HMI tags "DB_SDC_GLOBAL"
   "DB_SDC_GLOBAL_LIMITS[2].RAPID_SLOW" : Int = PLC DB_SDC_GLOBAL.LIMITS[2].RAPID_SLOW AT %DB3700.DBW512, 1 s   // Umstellung Begrenzung auf Abstand (mm), Einschränkung / Changeover limit of distance (mm), limitation
   "DB_SDC_GLOBAL_SYNCH[15].K" : Real = PLC DB_SDC_GLOBAL.SYNCH[15].K AT %DB3700.DBD426, 1 s   // erreichen von Synchron Faktor / gain for Synchron Faktor
   "DB_SDC_GLOBAL_SYNCH[15].SET_DIST" : Int = PLC DB_SDC_GLOBAL.SYNCH[15].SET_DIST AT %DB3700.DBW420, 1 s   // Set point value: distance (mm)
   "DB_SDC_GLOBAL_LIMITS[6].RAPID_SLOW" : Int = PLC DB_SDC_GLOBAL.LIMITS[6].RAPID_SLOW AT %DB3700.DBW536, 1 s   // Umstellung Begrenzung auf Abstand (mm), Einschränkung / Changeover limit of distance (mm), limitation
   "DB_SDC_GLOBAL_SYNCH[11].HYST" : Int = PLC DB_SDC_GLOBAL.SYNCH[11].HYST AT %DB3700.DBW352, 1 s   // IO Hysterese
   "DB_SDC_GLOBAL_SYNCH[6].MIN_FAKT" : Real = PLC DB_SDC_GLOBAL.SYNCH[6].MIN_FAKT AT %DB3700.DBD272, 1 s   // Faktor für minimale Synchronisiergeschwindigkeit / Faktor Speed for Synchron MIN
   "DB_SDC_GLOBAL_MIN_DIST_EMS[13]" : Int = PLC DB_SDC_GLOBAL.MIN_DIST_EMS[13] AT %DB3700.DBW126, 1 s   // minimum distance
   "DB_SDC_GLOBAL_SYNCH[8].MIN_FAKT" : Real = PLC DB_SDC_GLOBAL.SYNCH[8].MIN_FAKT AT %DB3700.DBD308, 1 s   // Faktor für minimale Synchronisiergeschwindigkeit / Faktor Speed for Synchron MIN
   "DB_SDC_GLOBAL_SYNCH[10].MIN_FAKT" : Real = PLC DB_SDC_GLOBAL.SYNCH[10].MIN_FAKT AT %DB3700.DBD344, 1 s   // Faktor für minimale Synchronisiergeschwindigkeit / Faktor Speed for Synchron MIN
   "DB_SDC_GLOBAL_SYNCH[6].SET_DIST" : Int = PLC DB_SDC_GLOBAL.SYNCH[6].SET_DIST AT %DB3700.DBW258, 1 s   // Set point value: distance (mm)
   "DB_SDC_GLOBAL_SYNCH[11].MAX_FAKT" : Real = PLC DB_SDC_GLOBAL.SYNCH[11].MAX_FAKT AT %DB3700.DBD358, 1 s   // Faktor für maximale Synchronisiergeschwindigkeit / Faktor Speed for Synchron MAX
   "DB_SDC_GLOBAL_SYNCH[9].SET_DIST" : Int = PLC DB_SDC_GLOBAL.SYNCH[9].SET_DIST AT %DB3700.DBW312, 1 s   // Set point value: distance (mm)
   "DB_SDC_GLOBAL_SYNCH[11].MIN_FAKT" : Real = PLC DB_SDC_GLOBAL.SYNCH[11].MIN_FAKT AT %DB3700.DBD362, 1 s   // Faktor für minimale Synchronisiergeschwindigkeit / Faktor Speed for Synchron MIN
   "DB_SDC_GLOBAL_MAN_V_1" : DInt = PLC DB_SDC_GLOBAL.MAN_V_1 AT %DB3700.DBD30, 1 s   // manual mode, set value: drive speed (mm/min)
   "DB_SDC_GLOBAL_LIMITS[5].RAPID_SLOW" : Int = PLC DB_SDC_GLOBAL.LIMITS[5].RAPID_SLOW AT %DB3700.DBW530, 1 s   // Umstellung Begrenzung auf Abstand (mm), Einschränkung / Changeover limit of distance (mm), limitation
   "DB_SDC_GLOBAL_SYNCH[13].MIN_FAKT" : Real = PLC DB_SDC_GLOBAL.SYNCH[13].MIN_FAKT AT %DB3700.DBD398, 1 s   // Faktor für minimale Synchronisiergeschwindigkeit / Faktor Speed for Synchron MIN
   "DB_SDC_GLOBAL_SYNCH[10].SET_DIST" : Int = PLC DB_SDC_GLOBAL.SYNCH[10].SET_DIST AT %DB3700.DBW330, 1 s   // Set point value: distance (mm)
   "DB_SDC_GLOBAL_SYNCH[9].HYST" : Int = PLC DB_SDC_GLOBAL.SYNCH[9].HYST AT %DB3700.DBW316, 1 s   // IO Hysterese
   "DB_SDC_GLOBAL_SYNCH[13].MAX_FAKT" : Real = PLC DB_SDC_GLOBAL.SYNCH[13].MAX_FAKT AT %DB3700.DBD394, 1 s   // Faktor für maximale Synchronisiergeschwindigkeit / Faktor Speed for Synchron MAX
   "DB_SDC_GLOBAL_LIMITS[11].RAPID_SLOW" : Int = PLC DB_SDC_GLOBAL.LIMITS[11].RAPID_SLOW AT %DB3700.DBW566, 1 s   // Umstellung Begrenzung auf Abstand (mm), Einschränkung / Changeover limit of distance (mm), limitation
   "DB_SDC_GLOBAL_SYNCH[3].MIN_FAKT" : Real = PLC DB_SDC_GLOBAL.SYNCH[3].MIN_FAKT AT %DB3700.DBD218, 1 s   // Faktor für minimale Synchronisiergeschwindigkeit / Faktor Speed for Synchron MIN
   "DB_SDC_GLOBAL_SYNCH[7].K" : Real = PLC DB_SDC_GLOBAL.SYNCH[7].K AT %DB3700.DBD282, 1 s   // erreichen von Synchron Faktor / gain for Synchron Faktor
   "DB_SDC_GLOBAL_SYNCH[2].SYNCH_DIST" : Int = PLC DB_SDC_GLOBAL.SYNCH[2].SYNCH_DIST AT %DB3700.DBW188, 1 s   // Start synchron distance value: distance (mm)
   "DB_SDC_GLOBAL_SYNCH[14].SYNCH_DIST" : Int = PLC DB_SDC_GLOBAL.SYNCH[14].SYNCH_DIST AT %DB3700.DBW404, 1 s   // Start synchron distance value: distance (mm)
   "DB_SDC_GLOBAL_MIN_DIST_EMS[8]" : Int = PLC DB_SDC_GLOBAL.MIN_DIST_EMS[8] AT %DB3700.DBW116, 1 s   // minimum distance
   "DB_SDC_GLOBAL_MIN_DIST_EMS[0]" : Int = PLC DB_SDC_GLOBAL.MIN_DIST_EMS[0] AT %DB3700.DBW100, 1 s   // minimum distance
   "DB_SDC_GLOBAL_SYNCH[14].K" : Real = PLC DB_SDC_GLOBAL.SYNCH[14].K AT %DB3700.DBD408, 1 s   // erreichen von Synchron Faktor / gain for Synchron Faktor
   "DB_SDC_GLOBAL_LIMITS[1].RAPID_SLOW" : Int = PLC DB_SDC_GLOBAL.LIMITS[1].RAPID_SLOW AT %DB3700.DBW506, 1 s   // Umstellung Begrenzung auf Abstand (mm), Einschränkung / Changeover limit of distance (mm), limitation
   "DB_SDC_GLOBAL_LIMITS[14].SLOW_SPEED_FAKT" : Real = PLC DB_SDC_GLOBAL.LIMITS[14].SLOW_SPEED_FAKT AT %DB3700.DBD586, 1 s   // Faktor Geschwindigkeit für langsame Drehzahl / Faktor Speed for Slow Speed
   "DB_SDC_GLOBAL_SYNCH[14].SET_DIST" : Int = PLC DB_SDC_GLOBAL.SYNCH[14].SET_DIST AT %DB3700.DBW402, 1 s   // Set point value: distance (mm)
   "DB_SDC_GLOBAL_SYNCH[15].SYNCH_DIST" : Int = PLC DB_SDC_GLOBAL.SYNCH[15].SYNCH_DIST AT %DB3700.DBW422, 1 s   // Start synchron distance value: distance (mm)
   "DB_SDC_GLOBAL_SYNCH[4].MAX_FAKT" : Real = PLC DB_SDC_GLOBAL.SYNCH[4].MAX_FAKT AT %DB3700.DBD232, 1 s   // Faktor für maximale Synchronisiergeschwindigkeit / Faktor Speed for Synchron MAX
   "DB_SDC_GLOBAL_SYNCH[2].HYST" : Int = PLC DB_SDC_GLOBAL.SYNCH[2].HYST AT %DB3700.DBW190, 1 s   // IO Hysterese
   "DB_SDC_GLOBAL_MIN_DIST_EMS[6]" : Int = PLC DB_SDC_GLOBAL.MIN_DIST_EMS[6] AT %DB3700.DBW112, 1 s   // minimum distance
   "DB_SDC_GLOBAL_SYNCH[0].HYST" : Int = PLC DB_SDC_GLOBAL.SYNCH[0].HYST AT %DB3700.DBW154, 1 s   // IO Hysterese
   "DB_SDC_GLOBAL_MIN_DIST_EMS[2]" : Int = PLC DB_SDC_GLOBAL.MIN_DIST_EMS[2] AT %DB3700.DBW104, 1 s   // minimum distance
   "DB_SDC_GLOBAL_MIN_DIST_EMS[12]" : Int = PLC DB_SDC_GLOBAL.MIN_DIST_EMS[12] AT %DB3700.DBW124, 1 s   // minimum distance
   "DB_SDC_GLOBAL_LIMITS[15].RAPID_SLOW" : Int = PLC DB_SDC_GLOBAL.LIMITS[15].RAPID_SLOW AT %DB3700.DBW590, 1 s   // Umstellung Begrenzung auf Abstand (mm), Einschränkung / Changeover limit of distance (mm), limitation
   "DB_SDC_GLOBAL_LIMITS[2].SLOW_SPEED_FAKT" : Real = PLC DB_SDC_GLOBAL.LIMITS[2].SLOW_SPEED_FAKT AT %DB3700.DBD514, 1 s   // Faktor Geschwindigkeit für langsame Drehzahl / Faktor Speed for Slow Speed
   "DB_SDC_GLOBAL_SYNCH[8].SET_DIST" : Int = PLC DB_SDC_GLOBAL.SYNCH[8].SET_DIST AT %DB3700.DBW294, 1 s   // Set point value: distance (mm)
   "DB_SDC_GLOBAL_min_barcode_mm" : DInt = PLC DB_SDC_GLOBAL.min_barcode_mm AT %DB3700.DBD6, 1 s   // Lower limit, bar code value
   "DB_SDC_GLOBAL_LIMITS[13].SLOW_SPEED_FAKT" : Real = PLC DB_SDC_GLOBAL.LIMITS[13].SLOW_SPEED_FAKT AT %DB3700.DBD580, 1 s   // Faktor Geschwindigkeit für langsame Drehzahl / Faktor Speed for Slow Speed
   "DB_SDC_GLOBAL_LIMITS[9].SLOW_SPEED_FAKT" : Real = PLC DB_SDC_GLOBAL.LIMITS[9].SLOW_SPEED_FAKT AT %DB3700.DBD556, 1 s   // Faktor Geschwindigkeit für langsame Drehzahl / Faktor Speed for Slow Speed
   "DB_SDC_GLOBAL_MIN_DIST_EMS[3]" : Int = PLC DB_SDC_GLOBAL.MIN_DIST_EMS[3] AT %DB3700.DBW106, 1 s   // minimum distance
   "DB_SDC_GLOBAL_SYNCH[4].SET_DIST" : Int = PLC DB_SDC_GLOBAL.SYNCH[4].SET_DIST AT %DB3700.DBW222, 1 s   // Set point value: distance (mm)
   "DB_SDC_GLOBAL_MAN_V_2" : DInt = PLC DB_SDC_GLOBAL.MAN_V_2 AT %DB3700.DBD34, 1 s   // manual mode, set value: drive speed (mm/min)
   "DB_SDC_GLOBAL_SYNCH[6].K" : Real = PLC DB_SDC_GLOBAL.SYNCH[6].K AT %DB3700.DBD264, 1 s   // erreichen von Synchron Faktor / gain for Synchron Faktor
   "DB_SDC_GLOBAL_SYNCH[2].K" : Real = PLC DB_SDC_GLOBAL.SYNCH[2].K AT %DB3700.DBD192, 1 s   // erreichen von Synchron Faktor / gain for Synchron Faktor
   "DB_SDC_GLOBAL_SYNCH[4].MIN_FAKT" : Real = PLC DB_SDC_GLOBAL.SYNCH[4].MIN_FAKT AT %DB3700.DBD236, 1 s   // Faktor für minimale Synchronisiergeschwindigkeit / Faktor Speed for Synchron MIN
   "DB_SDC_GLOBAL_SYNCH[6].SYNCH_DIST" : Int = PLC DB_SDC_GLOBAL.SYNCH[6].SYNCH_DIST AT %DB3700.DBW260, 1 s   // Start synchron distance value: distance (mm)
   "DB_SDC_GLOBAL_LIMITS[8].RAPID_SLOW" : Int = PLC DB_SDC_GLOBAL.LIMITS[8].RAPID_SLOW AT %DB3700.DBW548, 1 s   // Umstellung Begrenzung auf Abstand (mm), Einschränkung / Changeover limit of distance (mm), limitation
   "DB_SDC_GLOBAL_SYNCH[11].SET_DIST" : Int = PLC DB_SDC_GLOBAL.SYNCH[11].SET_DIST AT %DB3700.DBW348, 1 s   // Set point value: distance (mm)
   "DB_SDC_GLOBAL_SYNCH[15].HYST" : Int = PLC DB_SDC_GLOBAL.SYNCH[15].HYST AT %DB3700.DBW424, 1 s   // IO Hysterese
   "DB_SDC_GLOBAL_SYNCH[13].HYST" : Int = PLC DB_SDC_ERRORS_STAT.ER_AKT[50].ER_STAT[2].ERROR AT %DB3700.DBW388, 1 s   // IO Hysterese
   "DB_SDC_GLOBAL_SYNCH[5].MAX_FAKT" : Real = PLC DB_SDC_GLOBAL.SYNCH[5].MAX_FAKT AT %DB3700.DBD250, 1 s   // Faktor für maximale Synchronisiergeschwindigkeit / Faktor Speed for Synchron MAX
   "DB_SDC_GLOBAL_EMS_ID_MIN" : Int = PLC DB_SDC_GLOBAL.EMS_ID_MIN AT %DB3700.DBW2, 1 s   // Minimum EMS ID
   "DB_SDC_GLOBAL_SYNCH[5].K" : Real = PLC DB_SDC_GLOBAL.SYNCH[5].K AT %DB3700.DBD246, 1 s   // erreichen von Synchron Faktor / gain for Synchron Faktor
   "DB_SDC_GLOBAL_SYNCH[5].SET_DIST" : Int = PLC DB_SDC_GLOBAL.SYNCH[5].SET_DIST AT %DB3700.DBW240, 1 s   // Set point value: distance (mm)
   "DB_SDC_GLOBAL_SYNCH[0].SYNCH_DIST" : Int = PLC DB_SDC_GLOBAL.SYNCH[0].SYNCH_DIST AT %DB3700.DBW152, 1 s   // Start synchron distance value: distance (mm)
   "DB_SDC_GLOBAL_MIN_DIST_EMS[1]" : Int = PLC DB_SDC_GLOBAL.MIN_DIST_EMS[1] AT %DB3700.DBW102, 1 s   // minimum distance
   "DB_SDC_GLOBAL_SEK_MIN" : Int = PLC DB_SDC_GLOBAL.SEK_MIN AT %DB3700.DBW22, 1 s   // Erste Abschnitt Nummer / first section number
   "DB_SDC_GLOBAL_SYNCH[2].MAX_FAKT" : Real = PLC DB_SDC_GLOBAL.SYNCH[2].MAX_FAKT AT %DB3700.DBD196, 1 s   // Faktor für maximale Synchronisiergeschwindigkeit / Faktor Speed for Synchron MAX
   "DB_SDC_GLOBAL_SYNCH[1].MIN_FAKT" : Real = PLC DB_SDC_GLOBAL.SYNCH[1].MIN_FAKT AT %DB3700.DBD182, 1 s   // Faktor für minimale Synchronisiergeschwindigkeit / Faktor Speed for Synchron MIN
   "DB_SDC_GLOBAL_SYNCH[2].MIN_FAKT" : Real = PLC DB_SDC_GLOBAL.SYNCH[2].MIN_FAKT AT %DB3700.DBD200, 1 s   // Faktor für minimale Synchronisiergeschwindigkeit / Faktor Speed for Synchron MIN
   "DB_SDC_GLOBAL_LIMITS[10].RAPID_SLOW" : Int = PLC DB_SDC_GLOBAL.LIMITS[10].RAPID_SLOW AT %DB3700.DBW560, 1 s   // Umstellung Begrenzung auf Abstand (mm), Einschränkung / Changeover limit of distance (mm), limitation
   "DB_SDC_GLOBAL_SYNCH[6].MAX_FAKT" : Real = PLC DB_SDC_GLOBAL.SYNCH[6].MAX_FAKT AT %DB3700.DBD268, 1 s   // Faktor für maximale Synchronisiergeschwindigkeit / Faktor Speed for Synchron MAX
   "DB_SDC_GLOBAL_SYNCH[10].K" : Real = PLC DB_SDC_GLOBAL.SYNCH[10].K AT %DB3700.DBD336, 1 s   // erreichen von Synchron Faktor / gain for Synchron Faktor
   "DB_SDC_GLOBAL_END_COURSE" : DInt = PLC DB_SDC_GLOBAL.END_COURSE AT %DB3700.DBD18, 1 s   // Ende Barcodewert vom Kurs / End Barcodevalue of Course
   "DB_SDC_GLOBAL_SYNCH[1].SYNCH_DIST" : Int = PLC DB_SDC_GLOBAL.SYNCH[1].SYNCH_DIST AT %DB3700.DBW170, 1 s   // Start synchron distance value: distance (mm)
   "DB_SDC_GLOBAL_LIMITS[1].SLOW_SPEED_FAKT" : Real = PLC DB_SDC_GLOBAL.LIMITS[1].SLOW_SPEED_FAKT AT %DB3700.DBD508, 1 s   // Faktor Geschwindigkeit für langsame Drehzahl / Faktor Speed for Slow Speed
   "DB_SDC_GLOBAL_SYNCH[11].SYNCH_DIST" : Int = PLC DB_SDC_GLOBAL.SYNCH[11].SYNCH_DIST AT %DB3700.DBW350, 1 s   // Start synchron distance value: distance (mm)
   "DB_SDC_GLOBAL_SYNCH[12].HYST" : Int = PLC DB_SDC_GLOBAL.SYNCH[12].HYST AT %DB3700.DBW370, 1 s   // IO Hysterese
   "DB_SDC_GLOBAL_LIMITS[0].RAPID_SLOW" : Int = PLC DB_SDC_GLOBAL.LIMITS[0].RAPID_SLOW AT %DB3700.DBW500, 1 s   // Umstellung Begrenzung auf Abstand (mm), Einschränkung / Changeover limit of distance (mm), limitation
   "DB_SDC_GLOBAL_SYNCH[15].MIN_FAKT" : Real = PLC DB_SDC_GLOBAL.SYNCH[15].MIN_FAKT AT %DB3700.DBD434, 1 s   // Faktor für minimale Synchronisiergeschwindigkeit / Faktor Speed for Synchron MIN
   "DB_SDC_GLOBAL_LIMITS[11].SLOW_SPEED_FAKT" : Real = PLC DB_SDC_GLOBAL.LIMITS[11].SLOW_SPEED_FAKT AT %DB3700.DBD568, 1 s   // Faktor Geschwindigkeit für langsame Drehzahl / Faktor Speed for Slow Speed
   "DB_SDC_GLOBAL_LIMITS[6].SLOW_SPEED_FAKT" : Real = PLC DB_SDC_GLOBAL.LIMITS[6].SLOW_SPEED_FAKT AT %DB3700.DBD538, 1 s   // Faktor Geschwindigkeit für langsame Drehzahl / Faktor Speed for Slow Speed
   "DB_SDC_GLOBAL_SYNCH[3].SYNCH_DIST" : Int = PLC DB_SDC_GLOBAL.SYNCH[3].SYNCH_DIST AT %DB3700.DBW206, 1 s   // Start synchron distance value: distance (mm)
   "DB_SDC_GLOBAL_MIN_DIST_EMS[11]" : Int = PLC DB_SDC_GLOBAL.MIN_DIST_EMS[11] AT %DB3700.DBW122, 1 s   // minimum distance
   "DB_SDC_GLOBAL_SYNCH[9].MAX_FAKT" : Real = PLC DB_SDC_GLOBAL.SYNCH[9].MAX_FAKT AT %DB3700.DBD322, 1 s   // Faktor für maximale Synchronisiergeschwindigkeit / Faktor Speed for Synchron MAX
   "DB_SDC_GLOBAL_MIN_DIST_EMS[9]" : Int = PLC DB_SDC_GLOBAL.MIN_DIST_EMS[9] AT %DB3700.DBW118, 1 s   // minimum distance
   "DB_SDC_GLOBAL_LIMITS[0].SLOW_SPEED_FAKT" : Real = PLC DB_SDC_GLOBAL.LIMITS[0].SLOW_SPEED_FAKT AT %DB3700.DBD502, 1 s   // Faktor Geschwindigkeit für langsame Drehzahl / Faktor Speed for Slow Speed
   "DB_SDC_GLOBAL_SYNCH[7].MAX_FAKT" : Real = PLC DB_SDC_GLOBAL.SYNCH[7].MAX_FAKT AT %DB3700.DBD286, 1 s   // Faktor für maximale Synchronisiergeschwindigkeit / Faktor Speed for Synchron MAX
   "DB_SDC_GLOBAL_SYNCH[7].MIN_FAKT" : Real = PLC DB_SDC_GLOBAL.SYNCH[7].MIN_FAKT AT %DB3700.DBD290, 1 s   // Faktor für minimale Synchronisiergeschwindigkeit / Faktor Speed for Synchron MIN
   "DB_SDC_GLOBAL_SYNCH[1].MAX_FAKT" : Real = PLC DB_SDC_GLOBAL.SYNCH[1].MAX_FAKT AT %DB3700.DBD178, 1 s   // Faktor für maximale Synchronisiergeschwindigkeit / Faktor Speed for Synchron MAX
   "DB_SDC_GLOBAL_LIMITS[14].RAPID_SLOW" : Int = PLC DB_SDC_GLOBAL.LIMITS[14].RAPID_SLOW AT %DB3700.DBW584, 1 s   // Umstellung Begrenzung auf Abstand (mm), Einschränkung / Changeover limit of distance (mm), limitation
   "DB_SDC_GLOBAL_SYNCH[9].K" : Real = PLC DB_SDC_GLOBAL.SYNCH[9].K AT %DB3700.DBD318, 1 s   // erreichen von Synchron Faktor / gain for Synchron Faktor
   "DB_SDC_GLOBAL_LIMITS[12].SLOW_SPEED_FAKT" : Real = PLC DB_SDC_GLOBAL.LIMITS[12].SLOW_SPEED_FAKT AT %DB3700.DBD574, 1 s   // Faktor Geschwindigkeit für langsame Drehzahl / Faktor Speed for Slow Speed
   "DB_SDC_GLOBAL_SYNCH[10].SYNCH_DIST" : Int = PLC DB_SDC_GLOBAL.SYNCH[10].SYNCH_DIST AT %DB3700.DBW332, 1 s   // Start synchron distance value: distance (mm)
   "DB_SDC_GLOBAL_SYNCH[12].SET_DIST" : Int = PLC DB_SDC_GLOBAL.SYNCH[12].SET_DIST AT %DB3700.DBW366, 1 s   // Set point value: distance (mm)
   "DB_SDC_GLOBAL_SYNCH[4].SYNCH_DIST" : Int = PLC DB_SDC_GLOBAL.SYNCH[4].SYNCH_DIST AT %DB3700.DBW224, 1 s   // Start synchron distance value: distance (mm)
   "DB_SDC_GLOBAL_SYNCH[8].HYST" : Int = PLC DB_SDC_GLOBAL.SYNCH[8].HYST AT %DB3700.DBW298, 1 s   // IO Hysterese
   "DB_SDC_GLOBAL_SYNCH[11].K" : Real = PLC DB_SDC_GLOBAL.SYNCH[11].K AT %DB3700.DBD354, 1 s   // erreichen von Synchron Faktor / gain for Synchron Faktor
   "DB_SDC_GLOBAL_SYNCH[12].SYNCH_DIST" : Int = PLC DB_SDC_GLOBAL.SYNCH[12].SYNCH_DIST AT %DB3700.DBW368, 1 s   // Start synchron distance value: distance (mm)
   "DB_SDC_GLOBAL_LIMITS[15].SLOW_SPEED_FAKT" : Real = PLC DB_SDC_GLOBAL.LIMITS[15].SLOW_SPEED_FAKT AT %DB3700.DBD592, 1 s   // Faktor Geschwindigkeit für langsame Drehzahl / Faktor Speed for Slow Speed
   "DB_SDC_GLOBAL_MIN_DIST_EMS[14]" : Int = PLC DB_SDC_GLOBAL.MIN_DIST_EMS[14] AT %DB3700.DBW128, 1 s   // minimum distance
   "DB_SDC_GLOBAL_SYNCH[1].SET_DIST" : Int = PLC DB_SDC_GLOBAL.SYNCH[1].SET_DIST AT %DB3700.DBW168, 1 s   // Set point value: distance (mm)
   "DB_SDC_GLOBAL_SYNCH[1].HYST" : Int = PLC DB_SDC_GLOBAL.SYNCH[1].HYST AT %DB3700.DBW172, 1 s   // IO Hysterese
   "DB_SDC_GLOBAL_LIMITS[7].RAPID_SLOW" : Int = PLC DB_SDC_GLOBAL.LIMITS[7].RAPID_SLOW AT %DB3700.DBW542, 1 s   // Umstellung Begrenzung auf Abstand (mm), Einschränkung / Changeover limit of distance (mm), limitation
   "DB_SDC_GLOBAL_LIMITS[13].RAPID_SLOW" : Int = PLC DB_SDC_GLOBAL.LIMITS[13].RAPID_SLOW AT %DB3700.DBW578, 1 s   // Umstellung Begrenzung auf Abstand (mm), Einschränkung / Changeover limit of distance (mm), limitation
   "DB_SDC_GLOBAL_SYNCH[0].K" : Real = PLC DB_SDC_GLOBAL.SYNCH[0].K AT %DB3700.DBD156, 1 s   // erreichen von Synchron Faktor / gain for Synchron Faktor
   "DB_SDC_GLOBAL_LIMITS[12].RAPID_SLOW" : Int = PLC DB_SDC_GLOBAL.LIMITS[12].RAPID_SLOW AT %DB3700.DBW572, 1 s   // Umstellung Begrenzung auf Abstand (mm), Einschränkung / Changeover limit of distance (mm), limitation
   "DB_SDC_GLOBAL_SYNCH[1].K" : Real = PLC DB_SDC_GLOBAL.SYNCH[1].K AT %DB3700.DBD174, 1 s   // erreichen von Synchron Faktor / gain for Synchron Faktor
   "DB_SDC_GLOBAL_SYNCH[12].K" : Real = PLC DB_SDC_GLOBAL.SYNCH[12].K AT %DB3700.DBD372, 1 s   // erreichen von Synchron Faktor / gain for Synchron Faktor
   "DB_SDC_GLOBAL_SYNCH[7].SET_DIST" : Int = PLC DB_SDC_GLOBAL.SYNCH[7].SET_DIST AT %DB3700.DBW276, 1 s   // Set point value: distance (mm)
   "DB_SDC_GLOBAL_SYNCH[5].HYST" : Int = PLC DB_SDC_GLOBAL.SYNCH[5].HYST AT %DB3700.DBW244, 1 s   // IO Hysterese
   "DB_SDC_GLOBAL_MIN_DIST_EMS[7]" : Int = PLC DB_SDC_GLOBAL.MIN_DIST_EMS[7] AT %DB3700.DBW114, 1 s   // minimum distance
   "DB_SDC_GLOBAL_SYNCH[13].K" : Real = PLC DB_SDC_GLOBAL.SYNCH[13].K AT %DB3700.DBD390, 1 s   // erreichen von Synchron Faktor / gain for Synchron Faktor
   "DB_SDC_GLOBAL_SYNCH[14].MIN_FAKT" : Real = PLC DB_SDC_GLOBAL.SYNCH[14].MIN_FAKT AT %DB3700.DBD416, 1 s   // Faktor für minimale Synchronisiergeschwindigkeit / Faktor Speed for Synchron MIN
   "DB_SDC_GLOBAL_SYNCH[9].SYNCH_DIST" : Int = PLC DB_SDC_GLOBAL.SYNCH[9].SYNCH_DIST AT %DB3700.DBW314, 1 s   // Start synchron distance value: distance (mm)
   "DB_SDC_GLOBAL_SYNCH[5].MIN_FAKT" : Real = PLC DB_SDC_GLOBAL.SYNCH[5].MIN_FAKT AT %DB3700.DBD254, 1 s   // Faktor für minimale Synchronisiergeschwindigkeit / Faktor Speed for Synchron MIN
   "DB_SDC_GLOBAL_SYNCH[8].K" : Real = PLC DB_SDC_GLOBAL.SYNCH[8].K AT %DB3700.DBD300, 1 s   // erreichen von Synchron Faktor / gain for Synchron Faktor
   "DB_SDC_GLOBAL_LIMITS[3].SLOW_SPEED_FAKT" : Real = PLC DB_SDC_GLOBAL.LIMITS[3].SLOW_SPEED_FAKT AT %DB3700.DBD520, 1 s   // Faktor Geschwindigkeit für langsame Drehzahl / Faktor Speed for Slow Speed
   "DB_SDC_GLOBAL_SYNCH[4].HYST" : Int = PLC DB_SDC_GLOBAL.SYNCH[4].HYST AT %DB3700.DBW226, 1 s   // IO Hysterese
   "DB_SDC_GLOBAL_SYNCH[0].MIN_FAKT" : Real = PLC DB_SDC_GLOBAL.SYNCH[0].MIN_FAKT AT %DB3700.DBD164, 1 s   // Faktor für minimale Synchronisiergeschwindigkeit / Faktor Speed for Synchron MIN
   "DB_SDC_GLOBAL_MIN_DIST_EMS[5]" : Int = PLC DB_SDC_GLOBAL.MIN_DIST_EMS[5] AT %DB3700.DBW110, 1 s   // minimum distance
   "DB_SDC_GLOBAL_LIMITS[7].SLOW_SPEED_FAKT" : Real = PLC DB_SDC_GLOBAL.LIMITS[7].SLOW_SPEED_FAKT AT %DB3700.DBD544, 1 s   // Faktor Geschwindigkeit für langsame Drehzahl / Faktor Speed for Slow Speed
   "DB_SDC_GLOBAL_SEK_MAX" : Int = PLC DB_SDC_GLOBAL.SEK_MAX AT %DB3700.DBW24, 1 s   // Aktuelle Anzahl der Bahnabschnitte / Current quantity of track sections
   "DB_SDC_GLOBAL_SYNCH[8].MAX_FAKT" : Real = PLC DB_SDC_GLOBAL.SYNCH[8].MAX_FAKT AT %DB3700.DBD304, 1 s   // Faktor für maximale Synchronisiergeschwindigkeit / Faktor Speed for Synchron MAX
   "DB_SDC_GLOBAL_EMS_ID_MAX" : Int = PLC DB_SDC_GLOBAL.EMS_ID_MAX AT %DB3700.DBW4, 1 s   // Maximum EMS ID
   "DB_SDC_GLOBAL_SYNCH[9].MIN_FAKT" : Real = PLC DB_SDC_GLOBAL.SYNCH[9].MIN_FAKT AT %DB3700.DBD326, 1 s   // Faktor für minimale Synchronisiergeschwindigkeit / Faktor Speed for Synchron MIN
   "DB_SDC_GLOBAL_SYNCH[7].HYST" : Int = PLC DB_SDC_GLOBAL.SYNCH[7].HYST AT %DB3700.DBW280, 1 s   // IO Hysterese
   "DB_SDC_GLOBAL_EMS_ID_ACT" : Int = PLC DB_SDC_GLOBAL.EMS_ID_ACT AT %DB3700.DBW0, 1 s   // Aktuelle Anzahl der EMS-Treiber / Current quantity of EMS drivers
   "DB_SDC_GLOBAL_SYNCH[3].MAX_FAKT" : Real = PLC DB_SDC_GLOBAL.SYNCH[3].MAX_FAKT AT %DB3700.DBD214, 1 s   // Faktor für maximale Synchronisiergeschwindigkeit / Faktor Speed for Synchron MAX
   "DB_SDC_GLOBAL_SYNCH[13].SET_DIST" : Int = PLC DB_SDC_GLOBAL.SYNCH[13].SET_DIST AT %DB3700.DBW384, 1 s   // Set point value: distance (mm)
   "DB_SDC_GLOBAL_LIMITS[3].RAPID_SLOW" : Int = PLC DB_SDC_GLOBAL.LIMITS[3].RAPID_SLOW AT %DB3700.DBW518, 1 s   // Umstellung Begrenzung auf Abstand (mm), Einschränkung / Changeover limit of distance (mm), limitation
   "DB_SDC_GLOBAL_SYNCH[3].K" : Real = PLC DB_SDC_GLOBAL.SYNCH[3].K AT %DB3700.DBD210, 1 s   // erreichen von Synchron Faktor / gain for Synchron Faktor
   "DB_SDC_GLOBAL_SYNCH[13].SYNCH_DIST" : Int = PLC DB_SDC_GLOBAL.SYNCH[13].SYNCH_DIST AT %DB3700.DBW386, 1 s   // Start synchron distance value: distance (mm)
   "DB_SDC_GLOBAL_SYNCH[5].SYNCH_DIST" : Int = PLC DB_SDC_GLOBAL.SYNCH[5].SYNCH_DIST AT %DB3700.DBW242, 1 s   // Start synchron distance value: distance (mm)
   "DB_SDC_GLOBAL_SYNCH[6].HYST" : Int = PLC DB_SDC_GLOBAL.SYNCH[6].HYST AT %DB3700.DBW262, 1 s   // IO Hysterese
   "DB_SDC_GLOBAL_SYNCH[14].HYST" : Int = PLC DB_SDC_GLOBAL.SYNCH[14].HYST AT %DB3700.DBW406, 1 s   // IO Hysterese
   "DB_SDC_GLOBAL_START_COURSE" : DInt = PLC DB_SDC_GLOBAL.START_COURSE AT %DB3700.DBD14, 1 s   // Start Barcodevalue of Course
   "DB_SDC_GLOBAL_SYNCH[0].MAX_FAKT" : Real = PLC DB_SDC_GLOBAL.SYNCH[0].MAX_FAKT AT %DB3700.DBD160, 1 s   // Faktor für maximale Synchronisiergeschwindigkeit / Faktor Speed for Synchron MAX
   "DB_SDC_GLOBAL_SYNCH[2].SET_DIST" : Int = PLC DB_SDC_GLOBAL.SYNCH[2].SET_DIST AT %DB3700.DBW186, 1 s   // Set point value: distance (mm)
   "DB_SDC_GLOBAL_LIMITS[4].SLOW_SPEED_FAKT" : Real = PLC DB_SDC_GLOBAL.LIMITS[4].SLOW_SPEED_FAKT AT %DB3700.DBD526, 1 s   // Faktor Geschwindigkeit für langsame Drehzahl / Faktor Speed for Slow Speed
   "DB_SDC_GLOBAL_LIMITS[5].SLOW_SPEED_FAKT" : Real = PLC DB_SDC_GLOBAL.LIMITS[5].SLOW_SPEED_FAKT AT %DB3700.DBD532, 1 s   // Faktor Geschwindigkeit für langsame Drehzahl / Faktor Speed for Slow Speed
   "DB_SDC_GLOBAL_MIN_DIST_EMS[15]" : Int = PLC DB_SDC_GLOBAL.MIN_DIST_EMS[15] AT %DB3700.DBW130, 1 s   // minimum distance
   "DB_SDC_GLOBAL_SYNCH[12].MIN_FAKT" : Real = PLC DB_SDC_GLOBAL.SYNCH[12].MIN_FAKT AT %DB3700.DBD380, 1 s   // Faktor für minimale Synchronisiergeschwindigkeit / Faktor Speed for Synchron MIN
   "DB_SDC_GLOBAL_SYNCH[14].MAX_FAKT" : Real = PLC DB_SDC_GLOBAL.SYNCH[14].MAX_FAKT AT %DB3700.DBD412, 1 s   // Faktor für maximale Synchronisiergeschwindigkeit / Faktor Speed for Synchron MAX
   "DB_SDC_GLOBAL_SYNCH[10].MAX_FAKT" : Real = PLC DB_SDC_GLOBAL.SYNCH[10].MAX_FAKT AT %DB3700.DBD340, 1 s   // Faktor für maximale Synchronisiergeschwindigkeit / Faktor Speed for Synchron MAX
   "DB_SDC_GLOBAL_SYNCH[8].SYNCH_DIST" : Int = PLC DB_SDC_GLOBAL.SYNCH[8].SYNCH_DIST AT %DB3700.DBW296, 1 s   // Start synchron distance value: distance (mm)
   "DB_SDC_GLOBAL_max_barcode_mm" : DInt = PLC DB_SDC_GLOBAL.max_barcode_mm AT %DB3700.DBD10, 1 s   // Upper limit, bar code value
   "DB_SDC_GLOBAL_LIMITS[4].RAPID_SLOW" : Int = PLC DB_SDC_GLOBAL.LIMITS[4].RAPID_SLOW AT %DB3700.DBW524, 1 s   // Umstellung Begrenzung auf Abstand (mm), Einschränkung / Changeover limit of distance (mm), limitation
   "DB_SDC_GLOBAL_SYNCH[3].SET_DIST" : Int = PLC DB_SDC_GLOBAL.SYNCH[3].SET_DIST AT %DB3700.DBW204, 1 s   // Set point value: distance (mm)
   "DB_SDC_GLOBAL_SYNCH[10].HYST" : Int = PLC DB_SDC_GLOBAL.SYNCH[10].HYST AT %DB3700.DBW334, 1 s   // IO Hysterese
   "DB_SDC_GLOBAL_MIN_DIST_EMS[4]" : Int = PLC DB_SDC_GLOBAL.MIN_DIST_EMS[4] AT %DB3700.DBW108, 1 s   // minimum distance
   "DB_SDC_GLOBAL_SYNCH[7].SYNCH_DIST" : Int = PLC DB_SDC_GLOBAL.SYNCH[7].SYNCH_DIST AT %DB3700.DBW278, 1 s   // Start synchron distance value: distance (mm)
   "DB_SDC_GLOBAL_SYNCH[4].K" : Real = PLC DB_SDC_GLOBAL.SYNCH[4].K AT %DB3700.DBD228, 1 s   // erreichen von Synchron Faktor / gain for Synchron Faktor
   "DB_SDC_GLOBAL_SYNCH[0].SET_DIST" : Int = PLC DB_SDC_GLOBAL.SYNCH[0].SET_DIST AT %DB3700.DBW150, 1 s   // Set point value: distance (mm)
   "DB_SDC_GLOBAL_LIMITS[10].SLOW_SPEED_FAKT" : Real = PLC DB_SDC_GLOBAL.LIMITS[10].SLOW_SPEED_FAKT AT %DB3700.DBD562, 1 s   // Faktor Geschwindigkeit für langsame Drehzahl / Faktor Speed for Slow Speed
   "DB_SDC_GLOBAL_MIN_DIST_EMS[10]" : Int = PLC DB_SDC_GLOBAL.MIN_DIST_EMS[10] AT %DB3700.DBW120, 1 s   // minimum distance
   "DB_SDC_GLOBAL_SYNCH[15].MAX_FAKT" : Real = PLC DB_SDC_GLOBAL.SYNCH[15].MAX_FAKT AT %DB3700.DBD430, 1 s   // Faktor für maximale Synchronisiergeschwindigkeit / Faktor Speed for Synchron MAX
   "DB_SDC_GLOBAL_SYNCH[12].MAX_FAKT" : Real = PLC DB_SDC_GLOBAL.SYNCH[12].MAX_FAKT AT %DB3700.DBD376, 1 s   // Faktor für maximale Synchronisiergeschwindigkeit / Faktor Speed for Synchron MAX
   "DB_SDC_GLOBAL_LIMITS[8].SLOW_SPEED_FAKT" : Real = PLC DB_SDC_GLOBAL.LIMITS[8].SLOW_SPEED_FAKT AT %DB3700.DBD550, 1 s   // Faktor Geschwindigkeit für langsame Drehzahl / Faktor Speed for Slow Speed
   "DB_SDC_GLOBAL_LIMITS[9].RAPID_SLOW" : Int = PLC DB_SDC_GLOBAL.LIMITS[9].RAPID_SLOW AT %DB3700.DBW554, 1 s   // Umstellung Begrenzung auf Abstand (mm), Einschränkung / Changeover limit of distance (mm), limitation
   "DB_SDC_GLOBAL_SYNCH[3].HYST" : Int = PLC DB_SDC_GLOBAL.SYNCH[3].HYST AT %DB3700.DBW208, 1 s   // IO Hysterese
   "DB_SDC_GLOBAL_SEK_CYCLE_COUNTER" : Int = PLC DB_SDC_GLOBAL.SEK_CYCLE_COUNTER AT %DB3700.DBW28, 1 s
   "DB_SDC_GLOBAL_EMS_VCleaner_1" : Int = PLC DB_SDC_GLOBAL.EMS_VCleaner_1 AT %DB3700.DBW90, 1 s

HMI tags "DB_SDC_HMI"
   "DB_SDC_GLOBAL_M.SDC_ER_Reset(1)" : Bool = PLC DB_SDC_GLOBAL.M.SDC_ER_Reset AT %DB3700.DBX600.4, 1 s   // Fehler Reset / Fault Reset

HMI tags "VAT_DB_SDC_TS_REFERENCE"
   "DB_SDC_TS_REFERENCE_3_HEADER.MAX_NR_SEK" : Int = PLC DB_SDC_TS_REFERENCE_3.HEADER.MAX_NR_SEK AT %DB3782.DBW4, 1 s   // Höchste SEK Nummer im DB
   "DB_SDC_TS_REFERENCE_1_HEADER.MIN_NR_SEK" : Int = PLC DB_SDC_TS_REFERENCE_1.HEADER.MIN_NR_SEK AT %DB3780.DBW2, 1 s   // Niedrigste SEK Nummer im DB
   "SDC\DB_SDC_TS_REFERENCE\_TS_Ref_Byte_80" : DInt, internal
   "SDC\DB_SDC_TS_REFERENCE\DB_SDC_TS_REFERENCE_X.Reference[XXX].Hoist_offset_3" : Array [0..15] of Char AT %DB0.DBX0.0, 1 s   // definition Hub-Offset 3(mm)
   "DB_SDC_TS_REFERENCE_5_HEADER.MIN_NR_SEK" : Int = PLC DB_SDC_TS_REFERENCE_5.HEADER.MIN_NR_SEK AT %DB3784.DBW2, 1 s   // Niedrigste SEK Nummer im DB
   "DB_SDC_TS_REFERENCE_6_HEADER.DB_NR" : Int = PLC DB_SDC_TS_REFERENCE_6.HEADER.DB_NR AT %DB3785.DBW0, 1 s   // DB Nummer
   "DB_SDC_TS_REFERENCE_2_HEADER.DB_NR" : Int = PLC DB_SDC_TS_REFERENCE_2.HEADER.DB_NR AT %DB3781.DBW0, 1 s   // DB Nummer
   "SDC\DB_SDC_TS_REFERENCE\DB_SDC_TS_REFERENCE_X.Reference[XXX].Height" : Array [0..15] of Char AT %DB0.DBX0.0, 1 s   // definition Hubposition (mm)
   "DB_SDC_TS_REFERENCE_3_HEADER.DB_NR" : Int = PLC DB_SDC_TS_REFERENCE_3.HEADER.DB_NR AT %DB3782.DBW0, 1 s   // DB Nummer
   "DB_SDC_TS_REFERENCE_2_HEADER.MAX_NR_SEK" : Int = PLC DB_SDC_TS_REFERENCE_2.HEADER.MAX_NR_SEK AT %DB3781.DBW4, 1 s   // Höchste SEK Nummer im DB
   "SDC\DB_SDC_TS_REFERENCE\_TS_Ref_DB_Nr" : Int, internal
   "SDC\DB_SDC_TS_REFERENCE\DB_SDC_TS_REFERENCE_X.Reference[XXX].Sektion" : Array [0..15] of Char AT %DB0.DBX0.0, 1 s   // definition Sektion
   "DB_SDC_TS_REFERENCE_1_HEADER.MAX_NR_SEK" : Int = PLC DB_SDC_TS_REFERENCE_1.HEADER.MAX_NR_SEK AT %DB3780.DBW4, 1 s   // Höchste SEK Nummer im DB
   "SDC\DB_SDC_TS_REFERENCE\_TS_Ref_Byte_32" : DInt, internal
   "SDC\DB_SDC_TS_REFERENCE\_TS_Ref_Byte_64" : DInt, internal
   "DB_SDC_TS_REFERENCE_6_HEADER.MIN_NR_SEK" : Int = PLC DB_SDC_TS_REFERENCE_6.HEADER.MIN_NR_SEK AT %DB3785.DBW2, 1 s   // Niedrigste SEK Nummer im DB
   "SDC\DB_SDC_TS_REFERENCE\DB_SDC_TS_REFERENCE_X.Reference[XXX].Hoist_offset_4" : Array [0..15] of Char AT %DB0.DBX0.0, 1 s   // definition Hub-Offset 4 (mm)
   "DB_SDC_TS_REFERENCE_1_HEADER.DB_NR" : Int = PLC DB_SDC_TS_REFERENCE_1.HEADER.DB_NR AT %DB3780.DBW0, 1 s   // DB Nummer
   "SDC\DB_SDC_TS_REFERENCE\_TS_Ref_Byte_16" : DInt, internal
   "SDC\DB_SDC_TS_REFERENCE\_TS_Ref_Byte_00" : DInt, internal
   "SDC\DB_SDC_TS_REFERENCE\DB_SDC_TS_REFERENCE_X.Reference[XXX].Hoist_offset_1" : Array [0..15] of Char AT %DB0.DBX0.0, 1 s   // definition Hub-Offset 1 (mm)
   "SDC\DB_SDC_TS_REFERENCE\_TS_Ref_Byte_48" : DInt, internal
   "SDC\DB_SDC_TS_REFERENCE\_TS_Ref_Byte_96" : DInt, internal
   "DB_SDC_TS_REFERENCE_1_HEADER.START_DAT" : Int = PLC DB_SDC_TS_REFERENCE_1.HEADER.START_DAT AT %DB3780.DBW6, 1 s   // Startadresse der SEK im DB
   "DB_SDC_TS_REFERENCE_1_HEADER.LAENGE_SEK_DATA" : Int = PLC DB_SDC_TS_REFERENCE_1.HEADER.LAENGE_SEK_DATA AT %DB3780.DBW8, 1 s   // Länge SEK Data
   "SDC\DB_SDC_TS_REFERENCE\DB_SDC_TS_REFERENCE_X.Reference[XXX].Actionpoint_2" : Array [0..15] of Char AT %DB0.DBX0.0, 1 s   // definition Actionpoint 2
   "DB_SDC_TS_REFERENCE_4_HEADER.MIN_NR_SEK" : Int = PLC DB_SDC_TS_REFERENCE_4.HEADER.MIN_NR_SEK AT %DB3783.DBW2, 1 s   // Niedrigste SEK Nummer im DB
   "SDC\DB_SDC_TS_REFERENCE\DB_SDC_TS_REFERENCE_X.Reference[XXX].Actionpoint_1" : Array [0..15] of Char AT %DB0.DBX0.0, 1 s   // definition Actionpoint 1
   "DB_SDC_TS_REFERENCE_2_HEADER.MIN_NR_SEK" : Int = PLC DB_SDC_TS_REFERENCE_2.HEADER.MIN_NR_SEK AT %DB3781.DBW2, 1 s   // Niedrigste SEK Nummer im DB
   "DB_SDC_TS_REFERENCE_5_HEADER.DB_NR" : Int = PLC DB_SDC_TS_REFERENCE_5.HEADER.DB_NR AT %DB3784.DBW0, 1 s   // DB Nummer
   "SDC\DB_SDC_TS_REFERENCE\_TS_Ref_Byte_112" : DInt, internal
   "DB_SDC_TS_REFERENCE_5_HEADER.MAX_NR_SEK" : Int = PLC DB_SDC_TS_REFERENCE_5.HEADER.MAX_NR_SEK AT %DB3784.DBW4, 1 s   // Höchste SEK Nummer im DB
   "DB_SDC_TS_REFERENCE_4_HEADER.DB_NR" : Int = PLC DB_SDC_TS_REFERENCE_4.HEADER.DB_NR AT %DB3783.DBW0, 1 s   // DB Nummer
   "SDC\DB_SDC_TS_REFERENCE\_TS_Ref_Nr" : Int, internal
      on ChangeValue: "SDC_TS_REFERENCE"("SDC\_TS_Nr")
   "DB_SDC_TS_REFERENCE_3_HEADER.MIN_NR_SEK" : Int = PLC DB_SDC_TS_REFERENCE_3.HEADER.MIN_NR_SEK AT %DB3782.DBW2, 1 s   // Niedrigste SEK Nummer im DB
   "DB_SDC_TS_REFERENCE_4_HEADER.MAX_NR_SEK" : Int = PLC DB_SDC_TS_REFERENCE_4.HEADER.MAX_NR_SEK AT %DB3783.DBW4, 1 s   // Höchste SEK Nummer im DB
   "DB_SDC_TS_REFERENCE_6_HEADER.MAX_NR_SEK" : Int = PLC DB_SDC_TS_REFERENCE_6.HEADER.MAX_NR_SEK AT %DB3785.DBW4, 1 s   // Höchste SEK Nummer im DB
   "SDC\DB_SDC_TS_REFERENCE\DB_SDC_TS_REFERENCE_X.Reference[XXX].Hoist_offset_2" : Array [0..15] of Char AT %DB0.DBX0.0, 1 s   // definition Hub-Offset 2 (mm)
